REGION Network 10
   RUNG wire#powerrail
      Contact( "EstadosCmpALTA-MTA"._4s1 )
      I_Contact( "CompALTA-MTA".ReqMch4 )
      wire#w1
      Contact( "DB-CompAltaDatos".Aut4 )
      Coil( "Concatenadoras"._4c10 )
   END_RUNG
   RUNG wire#powerrail
      Contact( "EstadosCmpALTA-MTA"._4s9 )
      I_Contact( "CompALTA-MTA".ReqMch4 )
   END_RUNG wire#w1
   RUNG wire#powerrail
      Contact( "EstadosCmpALTA-MTA"._4s3 )
      I_Contact( "DB-CompAltaDatos".PanMchCmp4 )
   END_RUNG wire#w1
   // the same network as SCL:
   "Concatenadoras"._4c10 := (("EstadosCmpALTA-MTA"._4s1 AND NOT "CompALTA-MTA".ReqMch4) OR ("EstadosCmpALTA-MTA"._4s9 AND NOT "CompALTA-MTA".ReqMch4) OR ("EstadosCmpALTA-MTA"._4s3 AND NOT "DB-CompAltaDatos".PanMchCmp4)) AND "DB-CompAltaDatos".Aut4;
END_REGION

REGION Network 11
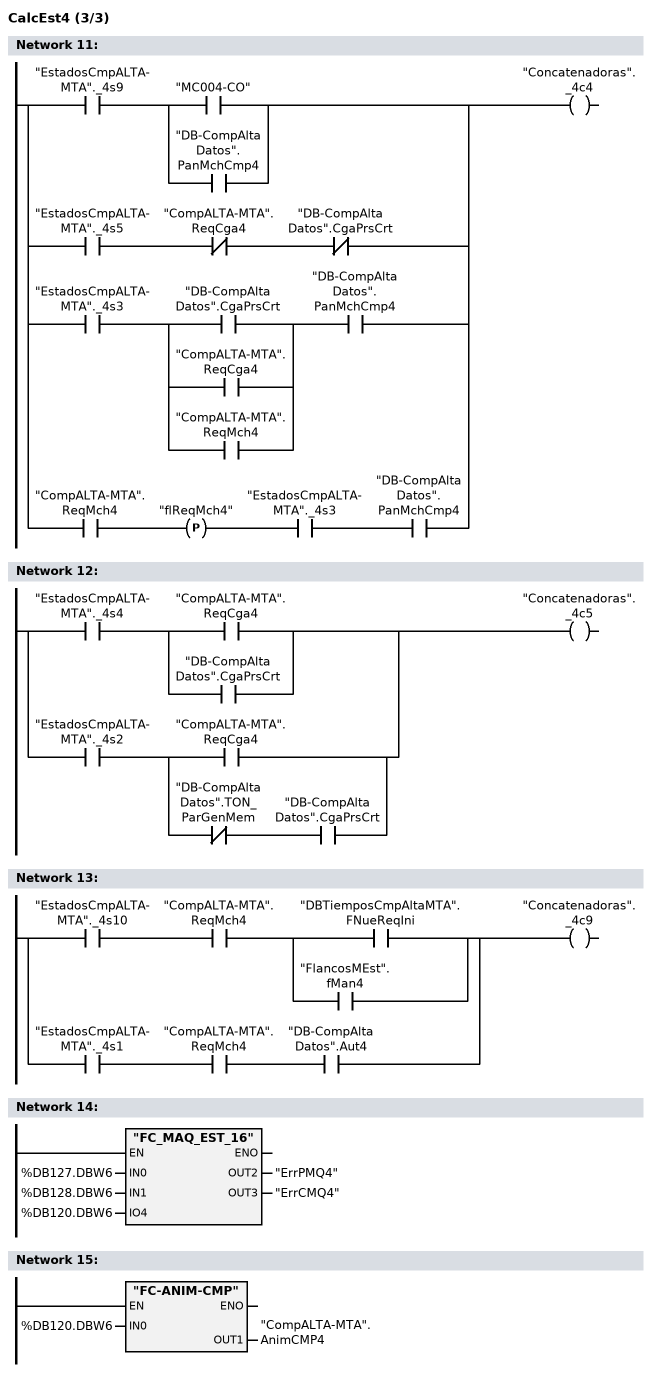
   RUNG wire#powerrail
      Contact( "EstadosCmpALTA-MTA"._4s9 )
      wire#w1
      Contact( "MC004-CO" )
      wire#w2
      Coil( "Concatenadoras"._4c4 )
   END_RUNG
   RUNG wire#w1
      Contact( "DB-CompAltaDatos".PanMchCmp4 )
   END_RUNG wire#w2
   RUNG wire#powerrail
      Contact( "EstadosCmpALTA-MTA"._4s5 )
      I_Contact( "CompALTA-MTA".ReqCga4 )
      I_Contact( "DB-CompAltaDatos".CgaPrsCrt )
   END_RUNG wire#w2
   RUNG wire#powerrail
      Contact( "EstadosCmpALTA-MTA"._4s3 )
      wire#w3
      Contact( "DB-CompAltaDatos".CgaPrsCrt )
      wire#w4
      Contact( "DB-CompAltaDatos".PanMchCmp4 )
   END_RUNG wire#w2
   RUNG wire#w3
      Contact( "CompALTA-MTA".ReqCga4 )
   END_RUNG wire#w4
   RUNG wire#w3
      Contact( "CompALTA-MTA".ReqMch4 )
   END_RUNG wire#w4
   RUNG wire#powerrail
      Contact( "CompALTA-MTA".ReqMch4 )
      P_Trig( "flReqMch4" )
      Contact( "EstadosCmpALTA-MTA"._4s3 )
      Contact( "DB-CompAltaDatos".PanMchCmp4 )
   END_RUNG wire#w2
   // the same network as SCL:
   #_w1 := "CompALTA-MTA".ReqMch4 AND NOT "flReqMch4";   // rising edge
   "flReqMch4" := "CompALTA-MTA".ReqMch4;
   "Concatenadoras"._4c4 := ("EstadosCmpALTA-MTA"._4s9 AND ("MC004-CO" OR "DB-CompAltaDatos".PanMchCmp4)) OR ("EstadosCmpALTA-MTA"._4s5 AND NOT "CompALTA-MTA".ReqCga4 AND NOT "DB-CompAltaDatos".CgaPrsCrt) OR ("EstadosCmpALTA-MTA"._4s3 AND ("DB-CompAltaDatos".CgaPrsCrt OR "CompALTA-MTA".ReqCga4 OR "CompALTA-MTA".ReqMch4) AND "DB-CompAltaDatos".PanMchCmp4) OR (#_w1 AND "EstadosCmpALTA-MTA"._4s3 AND "DB-CompAltaDatos".PanMchCmp4);
END_REGION

REGION Network 12
   RUNG wire#powerrail
      Contact( "EstadosCmpALTA-MTA"._4s4 )
      wire#w1
      Contact( "CompALTA-MTA".ReqCga4 )
      wire#w2
      Coil( "Concatenadoras"._4c5 )
   END_RUNG
   RUNG wire#w1
      Contact( "DB-CompAltaDatos".CgaPrsCrt )
   END_RUNG wire#w2
   RUNG wire#powerrail
      Contact( "EstadosCmpALTA-MTA"._4s2 )
      wire#w3
      Contact( "CompALTA-MTA".ReqCga4 )
   END_RUNG wire#w2
   RUNG wire#w3
      I_Contact( "DB-CompAltaDatos".TON_ParGenMem )
      Contact( "DB-CompAltaDatos".CgaPrsCrt )
   END_RUNG wire#w2
   // the same network as SCL:
   "Concatenadoras"._4c5 := ("EstadosCmpALTA-MTA"._4s4 AND ("CompALTA-MTA".ReqCga4 OR "DB-CompAltaDatos".CgaPrsCrt)) OR ("EstadosCmpALTA-MTA"._4s2 AND ("CompALTA-MTA".ReqCga4 OR (NOT "DB-CompAltaDatos".TON_ParGenMem AND "DB-CompAltaDatos".CgaPrsCrt)));
END_REGION

REGION Network 13
   RUNG wire#powerrail
      Contact( "EstadosCmpALTA-MTA"._4s10 )
      Contact( "CompALTA-MTA".ReqMch4 )
      wire#w1
      Contact( "DBTiemposCmpAltaMTA".FNueReqIni )
      wire#w2
      Coil( "Concatenadoras"._4c9 )
   END_RUNG
   RUNG wire#w1
      Contact( "FlancosMEst".fMan4 )
   END_RUNG wire#w2
   RUNG wire#powerrail
      Contact( "EstadosCmpALTA-MTA"._4s1 )
      Contact( "CompALTA-MTA".ReqMch4 )
      Contact( "DB-CompAltaDatos".Aut4 )
   END_RUNG wire#w2
   // the same network as SCL:
   "Concatenadoras"._4c9 := ("EstadosCmpALTA-MTA"._4s10 AND "CompALTA-MTA".ReqMch4 AND ("DBTiemposCmpAltaMTA".FNueReqIni OR "FlancosMEst".fMan4)) OR ("EstadosCmpALTA-MTA"._4s1 AND "CompALTA-MTA".ReqMch4 AND "DB-CompAltaDatos".Aut4);
END_REGION

REGION Network 14
   RUNG wire#powerrail
      "FC_MAQ_EST_16"(IN0 := %DB127.DBW6, IN1 := %DB128.DBW6, IO4 := %DB120.DBW6, OUT2 => "ErrPMQ4", OUT3 => "ErrCMQ4")
   END_RUNG
   // the same network as SCL:
   "FC_MAQ_EST_16"(IN0 := %DB127.DBW6,
                   IN1 := %DB128.DBW6,
                   IO4 := %DB120.DBW6,
                   OUT2 => "ErrPMQ4",
                   OUT3 => "ErrCMQ4");
END_REGION

REGION Network 15
   RUNG wire#powerrail
      "FC-ANIM-CMP"(IN0 := %DB120.DBW6, OUT1 => "CompALTA-MTA".AnimCMP4)
   END_RUNG
   // the same network as SCL:
   "FC-ANIM-CMP"(IN0 := %DB120.DBW6, OUT1 => "CompALTA-MTA".AnimCMP4);
END_REGION
END_FUNCTION

FUNCTION "CalcEst5" : Void   // FC40, LAD
{ S7_Optimized_Access := 'FALSE' }
VERSION : 0.1
   VAR_TEMP   // added for the SCL form of the ladder/FBD networks
      _w1 : Bool;
   END_VAR
BEGIN

REGION Network 1: Prioritaria 1
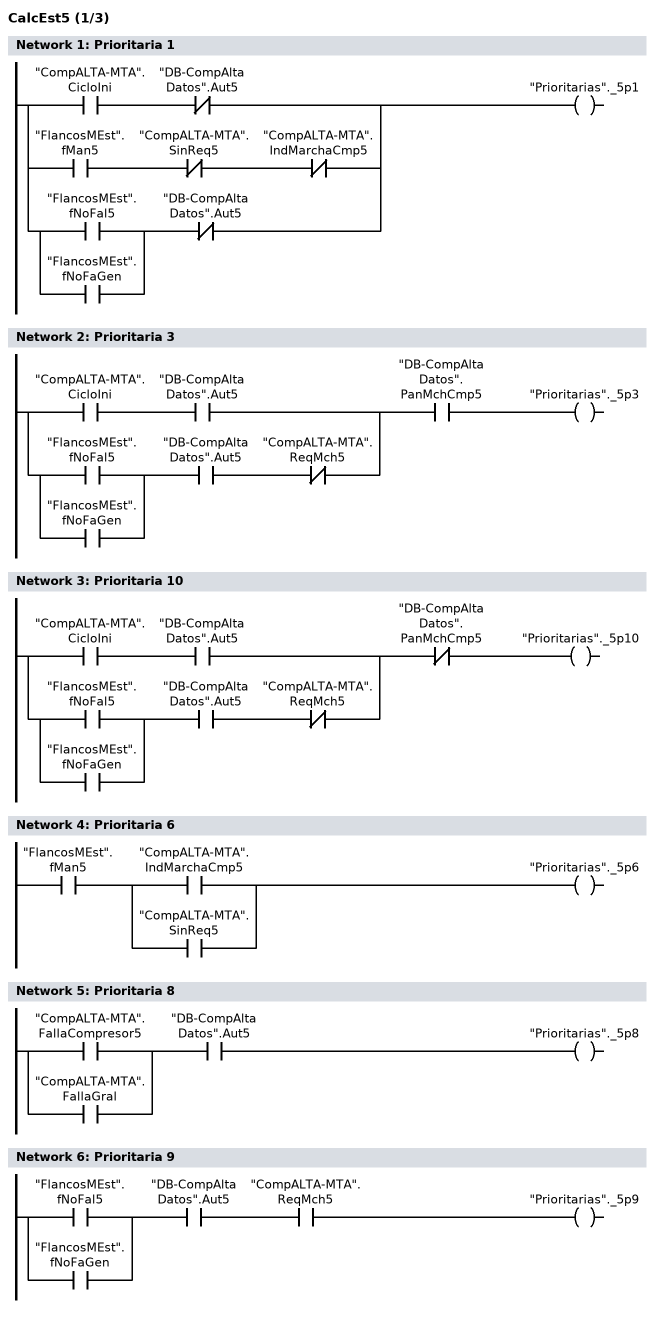
   RUNG wire#powerrail
      Contact( "CompALTA-MTA".CicloIni )
      I_Contact( "DB-CompAltaDatos".Aut5 )
      wire#w1
      Coil( "Prioritarias"._5p1 )
   END_RUNG
   RUNG wire#powerrail
      Contact( "FlancosMEst".fMan5 )
      I_Contact( "CompALTA-MTA".SinReq5 )
      I_Contact( "CompALTA-MTA".IndMarchaCmp5 )
   END_RUNG wire#w1
   RUNG wire#powerrail
      Contact( "FlancosMEst".fNoFal5 )
      wire#w2
      I_Contact( "DB-CompAltaDatos".Aut5 )
   END_RUNG wire#w1
   RUNG wire#powerrail
      Contact( "FlancosMEst".fNoFaGen )
   END_RUNG wire#w2
   // the same network as SCL:
   "Prioritarias"._5p1 := ("CompALTA-MTA".CicloIni AND NOT "DB-CompAltaDatos".Aut5) OR ("FlancosMEst".fMan5 AND NOT "CompALTA-MTA".SinReq5 AND NOT "CompALTA-MTA".IndMarchaCmp5) OR (("FlancosMEst".fNoFal5 OR "FlancosMEst".fNoFaGen) AND NOT "DB-CompAltaDatos".Aut5);
END_REGION

REGION Network 2: Prioritaria 3
   RUNG wire#powerrail
      Contact( "CompALTA-MTA".CicloIni )
      Contact( "DB-CompAltaDatos".Aut5 )
      wire#w1
      Contact( "DB-CompAltaDatos".PanMchCmp5 )
      Coil( "Prioritarias"._5p3 )
   END_RUNG
   RUNG wire#powerrail
      Contact( "FlancosMEst".fNoFal5 )
      wire#w2
      Contact( "DB-CompAltaDatos".Aut5 )
      I_Contact( "CompALTA-MTA".ReqMch5 )
   END_RUNG wire#w1
   RUNG wire#powerrail
      Contact( "FlancosMEst".fNoFaGen )
   END_RUNG wire#w2
   // the same network as SCL:
   "Prioritarias"._5p3 := (("CompALTA-MTA".CicloIni AND "DB-CompAltaDatos".Aut5) OR (("FlancosMEst".fNoFal5 OR "FlancosMEst".fNoFaGen) AND "DB-CompAltaDatos".Aut5 AND NOT "CompALTA-MTA".ReqMch5)) AND "DB-CompAltaDatos".PanMchCmp5;
END_REGION

REGION Network 3: Prioritaria 10
   RUNG wire#powerrail
      Contact( "CompALTA-MTA".CicloIni )
      Contact( "DB-CompAltaDatos".Aut5 )
      wire#w1
      I_Contact( "DB-CompAltaDatos".PanMchCmp5 )
      Coil( "Prioritarias"._5p10 )
   END_RUNG
   RUNG wire#powerrail
      Contact( "FlancosMEst".fNoFal5 )
      wire#w2
      Contact( "DB-CompAltaDatos".Aut5 )
      I_Contact( "CompALTA-MTA".ReqMch5 )
   END_RUNG wire#w1
   RUNG wire#powerrail
      Contact( "FlancosMEst".fNoFaGen )
   END_RUNG wire#w2
   // the same network as SCL:
   "Prioritarias"._5p10 := (("CompALTA-MTA".CicloIni AND "DB-CompAltaDatos".Aut5) OR (("FlancosMEst".fNoFal5 OR "FlancosMEst".fNoFaGen) AND "DB-CompAltaDatos".Aut5 AND NOT "CompALTA-MTA".ReqMch5)) AND NOT "DB-CompAltaDatos".PanMchCmp5;
END_REGION

REGION Network 4: Prioritaria 6
   RUNG wire#powerrail
      Contact( "FlancosMEst".fMan5 )
      wire#w1
      Contact( "CompALTA-MTA".IndMarchaCmp5 )
      wire#w2
      Coil( "Prioritarias"._5p6 )
   END_RUNG
   RUNG wire#w1
      Contact( "CompALTA-MTA".SinReq5 )
   END_RUNG wire#w2
   // the same network as SCL:
   "Prioritarias"._5p6 := "FlancosMEst".fMan5 AND ("CompALTA-MTA".IndMarchaCmp5 OR "CompALTA-MTA".SinReq5);
END_REGION

REGION Network 5: Prioritaria 8
   RUNG wire#powerrail
      Contact( "CompALTA-MTA".FallaCompresor5 )
      wire#w1
      Contact( "DB-CompAltaDatos".Aut5 )
      Coil( "Prioritarias"._5p8 )
   END_RUNG
   RUNG wire#powerrail
      Contact( "CompALTA-MTA".FallaGral )
   END_RUNG wire#w1
   // the same network as SCL:
   "Prioritarias"._5p8 := ("CompALTA-MTA".FallaCompresor5 OR "CompALTA-MTA".FallaGral) AND "DB-CompAltaDatos".Aut5;
END_REGION

REGION Network 6: Prioritaria 9
   RUNG wire#powerrail
      Contact( "FlancosMEst".fNoFal5 )
      wire#w1
      Contact( "DB-CompAltaDatos".Aut5 )
      Contact( "CompALTA-MTA".ReqMch5 )
      Coil( "Prioritarias"._5p9 )
   END_RUNG
   RUNG wire#powerrail
      Contact( "FlancosMEst".fNoFaGen )
   END_RUNG wire#w1
   // the same network as SCL:
   "Prioritarias"._5p9 := ("FlancosMEst".fNoFal5 OR "FlancosMEst".fNoFaGen) AND "DB-CompAltaDatos".Aut5 AND "CompALTA-MTA".ReqMch5;
END_REGION

REGION Network 7: Concatenadora 1
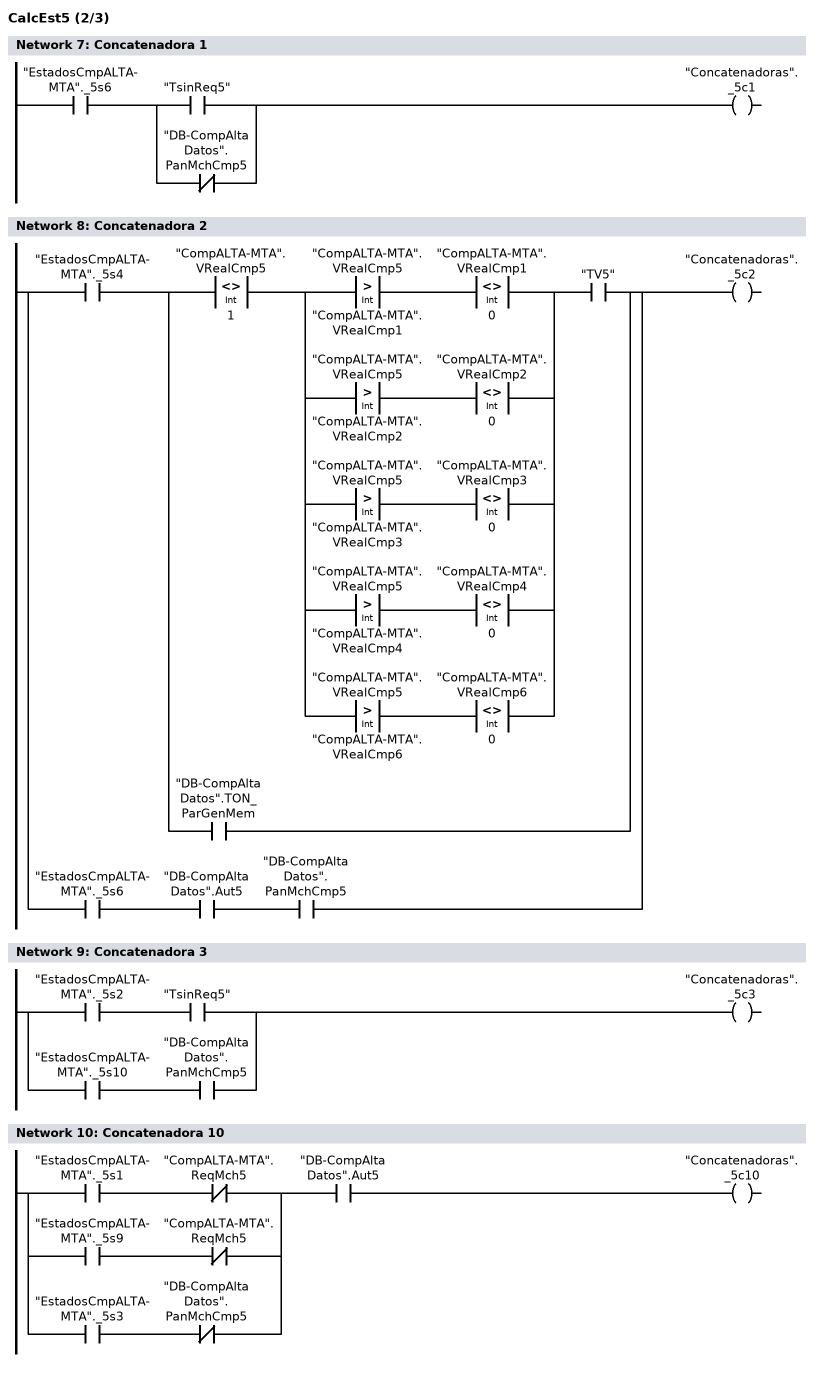
   RUNG wire#powerrail
      Contact( "EstadosCmpALTA-MTA"._5s6 )
      wire#w1
      Contact( "TsinReq5" )
      wire#w2
      Coil( "Concatenadoras"._5c1 )
   END_RUNG
   RUNG wire#w1
      I_Contact( "DB-CompAltaDatos".PanMchCmp5 )
   END_RUNG wire#w2
   // the same network as SCL:
   "Concatenadoras"._5c1 := "EstadosCmpALTA-MTA"._5s6 AND ("TsinReq5" OR NOT "DB-CompAltaDatos".PanMchCmp5);
END_REGION

REGION Network 8: Concatenadora 2
   RUNG wire#powerrail
      Contact( "EstadosCmpALTA-MTA"._5s4 )
      wire#w1
      { S7_Templates := "SrcType := Int" } NE_Contact(in1 := "CompALTA-MTA".VRealCmp5, in2 := 1)
      wire#w2
      { S7_Templates := "SrcType := Int" } GT_Contact(in1 := "CompALTA-MTA".VRealCmp5, in2 := "CompALTA-MTA".VRealCmp1)
      { S7_Templates := "SrcType := Int" } NE_Contact(in1 := "CompALTA-MTA".VRealCmp1, in2 := 0)
      wire#w3
      Contact( "TV5" )
      wire#w4
      Coil( "Concatenadoras"._5c2 )
   END_RUNG
   RUNG wire#w2
      { S7_Templates := "SrcType := Int" } GT_Contact(in1 := "CompALTA-MTA".VRealCmp5, in2 := "CompALTA-MTA".VRealCmp2)
      { S7_Templates := "SrcType := Int" } NE_Contact(in1 := "CompALTA-MTA".VRealCmp2, in2 := 0)
   END_RUNG wire#w3
   RUNG wire#w2
      { S7_Templates := "SrcType := Int" } GT_Contact(in1 := "CompALTA-MTA".VRealCmp5, in2 := "CompALTA-MTA".VRealCmp3)
      { S7_Templates := "SrcType := Int" } NE_Contact(in1 := "CompALTA-MTA".VRealCmp3, in2 := 0)
   END_RUNG wire#w3
   RUNG wire#w2
      { S7_Templates := "SrcType := Int" } GT_Contact(in1 := "CompALTA-MTA".VRealCmp5, in2 := "CompALTA-MTA".VRealCmp4)
      { S7_Templates := "SrcType := Int" } NE_Contact(in1 := "CompALTA-MTA".VRealCmp4, in2 := 0)
   END_RUNG wire#w3
   RUNG wire#w2
      { S7_Templates := "SrcType := Int" } GT_Contact(in1 := "CompALTA-MTA".VRealCmp5, in2 := "CompALTA-MTA".VRealCmp6)
      { S7_Templates := "SrcType := Int" } NE_Contact(in1 := "CompALTA-MTA".VRealCmp6, in2 := 0)
   END_RUNG wire#w3
   RUNG wire#w1
      Contact( "DB-CompAltaDatos".TON_ParGenMem )
   END_RUNG wire#w4
   RUNG wire#powerrail
      Contact( "EstadosCmpALTA-MTA"._5s6 )
      Contact( "DB-CompAltaDatos".Aut5 )
      Contact( "DB-CompAltaDatos".PanMchCmp5 )
   END_RUNG wire#w4
   // the same network as SCL:
   "Concatenadoras"._5c2 := ("EstadosCmpALTA-MTA"._5s4 AND ((("CompALTA-MTA".VRealCmp5 <> 1) AND ((("CompALTA-MTA".VRealCmp5 > "CompALTA-MTA".VRealCmp1) AND ("CompALTA-MTA".VRealCmp1 <> 0)) OR (("CompALTA-MTA".VRealCmp5 > "CompALTA-MTA".VRealCmp2) AND ("CompALTA-MTA".VRealCmp2 <> 0)) OR (("CompALTA-MTA".VRealCmp5 > "CompALTA-MTA".VRealCmp3) AND ("CompALTA-MTA".VRealCmp3 <> 0)) OR (("CompALTA-MTA".VRealCmp5 > "CompALTA-MTA".VRealCmp4) AND ("CompALTA-MTA".VRealCmp4 <> 0)) OR (("CompALTA-MTA".VRealCmp5 > "CompALTA-MTA".VRealCmp6) AND ("CompALTA-MTA".VRealCmp6 <> 0))) AND "TV5") OR "DB-CompAltaDatos".TON_ParGenMem)) OR ("EstadosCmpALTA-MTA"._5s6 AND "DB-CompAltaDatos".Aut5 AND "DB-CompAltaDatos".PanMchCmp5);
END_REGION

REGION Network 9: Concatenadora 3
   RUNG wire#powerrail
      Contact( "EstadosCmpALTA-MTA"._5s2 )
      Contact( "TsinReq5" )
      wire#w1
      Coil( "Concatenadoras"._5c3 )
   END_RUNG
   RUNG wire#powerrail
      Contact( "EstadosCmpALTA-MTA"._5s10 )
      Contact( "DB-CompAltaDatos".PanMchCmp5 )
   END_RUNG wire#w1
   // the same network as SCL:
   "Concatenadoras"._5c3 := ("EstadosCmpALTA-MTA"._5s2 AND "TsinReq5") OR ("EstadosCmpALTA-MTA"._5s10 AND "DB-CompAltaDatos".PanMchCmp5);
END_REGION

REGION Network 10: Concatenadora 10
   RUNG wire#powerrail
      Contact( "EstadosCmpALTA-MTA"._5s1 )
      I_Contact( "CompALTA-MTA".ReqMch5 )
      wire#w1
      Contact( "DB-CompAltaDatos".Aut5 )
      Coil( "Concatenadoras"._5c10 )
   END_RUNG
   RUNG wire#powerrail
      Contact( "EstadosCmpALTA-MTA"._5s9 )
      I_Contact( "CompALTA-MTA".ReqMch5 )
   END_RUNG wire#w1
   RUNG wire#powerrail
      Contact( "EstadosCmpALTA-MTA"._5s3 )
      I_Contact( "DB-CompAltaDatos".PanMchCmp5 )
   END_RUNG wire#w1
   // the same network as SCL:
   "Concatenadoras"._5c10 := (("EstadosCmpALTA-MTA"._5s1 AND NOT "CompALTA-MTA".ReqMch5) OR ("EstadosCmpALTA-MTA"._5s9 AND NOT "CompALTA-MTA".ReqMch5) OR ("EstadosCmpALTA-MTA"._5s3 AND NOT "DB-CompAltaDatos".PanMchCmp5)) AND "DB-CompAltaDatos".Aut5;
END_REGION

REGION Network 11: Concatenadora 4
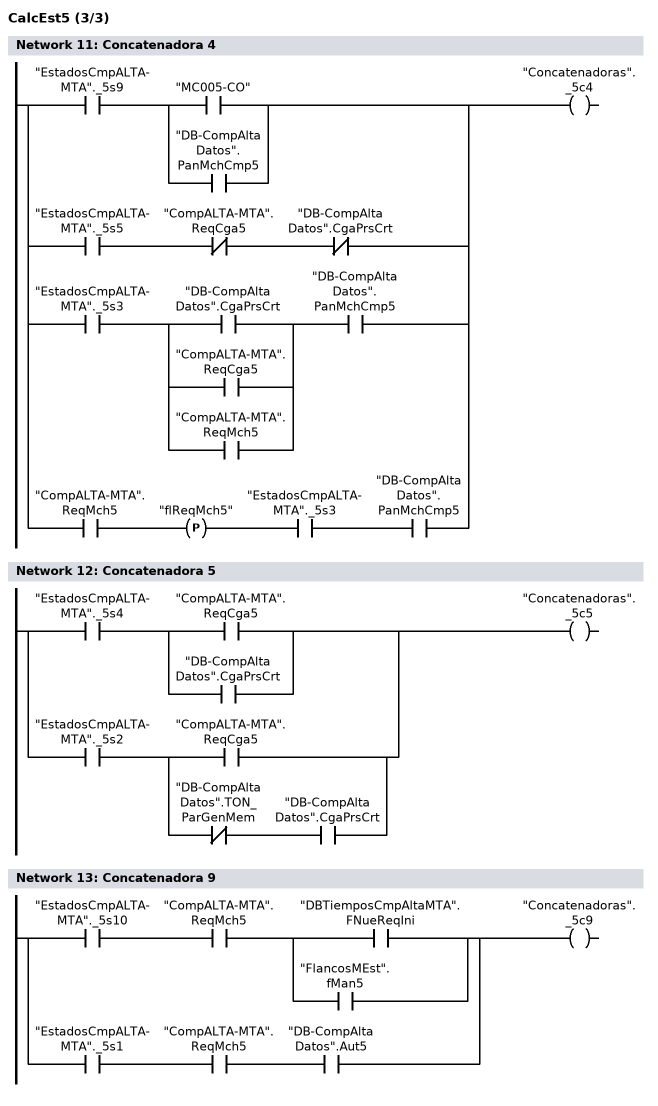
   RUNG wire#powerrail
      Contact( "EstadosCmpALTA-MTA"._5s9 )
      wire#w1
      Contact( "MC005-CO" )
      wire#w2
      Coil( "Concatenadoras"._5c4 )
   END_RUNG
   RUNG wire#w1
      Contact( "DB-CompAltaDatos".PanMchCmp5 )
   END_RUNG wire#w2
   RUNG wire#powerrail
      Contact( "EstadosCmpALTA-MTA"._5s5 )
      I_Contact( "CompALTA-MTA".ReqCga5 )
      I_Contact( "DB-CompAltaDatos".CgaPrsCrt )
   END_RUNG wire#w2
   RUNG wire#powerrail
      Contact( "EstadosCmpALTA-MTA"._5s3 )
      wire#w3
      Contact( "DB-CompAltaDatos".CgaPrsCrt )
      wire#w4
      Contact( "DB-CompAltaDatos".PanMchCmp5 )
   END_RUNG wire#w2
   RUNG wire#w3
      Contact( "CompALTA-MTA".ReqCga5 )
   END_RUNG wire#w4
   RUNG wire#w3
      Contact( "CompALTA-MTA".ReqMch5 )
   END_RUNG wire#w4
   RUNG wire#powerrail
      Contact( "CompALTA-MTA".ReqMch5 )
      P_Trig( "flReqMch5" )
      Contact( "EstadosCmpALTA-MTA"._5s3 )
      Contact( "DB-CompAltaDatos".PanMchCmp5 )
   END_RUNG wire#w2
   // the same network as SCL:
   #_w1 := "CompALTA-MTA".ReqMch5 AND NOT "flReqMch5";   // rising edge
   "flReqMch5" := "CompALTA-MTA".ReqMch5;
   "Concatenadoras"._5c4 := ("EstadosCmpALTA-MTA"._5s9 AND ("MC005-CO" OR "DB-CompAltaDatos".PanMchCmp5)) OR ("EstadosCmpALTA-MTA"._5s5 AND NOT "CompALTA-MTA".ReqCga5 AND NOT "DB-CompAltaDatos".CgaPrsCrt) OR ("EstadosCmpALTA-MTA"._5s3 AND ("DB-CompAltaDatos".CgaPrsCrt OR "CompALTA-MTA".ReqCga5 OR "CompALTA-MTA".ReqMch5) AND "DB-CompAltaDatos".PanMchCmp5) OR (#_w1 AND "EstadosCmpALTA-MTA"._5s3 AND "DB-CompAltaDatos".PanMchCmp5);
END_REGION

REGION Network 12: Concatenadora 5
   RUNG wire#powerrail
      Contact( "EstadosCmpALTA-MTA"._5s4 )
      wire#w1
      Contact( "CompALTA-MTA".ReqCga5 )
      wire#w2
      Coil( "Concatenadoras"._5c5 )
   END_RUNG
   RUNG wire#w1
      Contact( "DB-CompAltaDatos".CgaPrsCrt )
   END_RUNG wire#w2
   RUNG wire#powerrail
      Contact( "EstadosCmpALTA-MTA"._5s2 )
      wire#w3
      Contact( "CompALTA-MTA".ReqCga5 )
   END_RUNG wire#w2
   RUNG wire#w3
      I_Contact( "DB-CompAltaDatos".TON_ParGenMem )
      Contact( "DB-CompAltaDatos".CgaPrsCrt )
   END_RUNG wire#w2
   // the same network as SCL:
   "Concatenadoras"._5c5 := ("EstadosCmpALTA-MTA"._5s4 AND ("CompALTA-MTA".ReqCga5 OR "DB-CompAltaDatos".CgaPrsCrt)) OR ("EstadosCmpALTA-MTA"._5s2 AND ("CompALTA-MTA".ReqCga5 OR (NOT "DB-CompAltaDatos".TON_ParGenMem AND "DB-CompAltaDatos".CgaPrsCrt)));
END_REGION

REGION Network 13: Concatenadora 9
   RUNG wire#powerrail
      Contact( "EstadosCmpALTA-MTA"._5s10 )
      Contact( "CompALTA-MTA".ReqMch5 )
      wire#w1
      Contact( "DBTiemposCmpAltaMTA".FNueReqIni )
      wire#w2
      Coil( "Concatenadoras"._5c9 )
   END_RUNG
   RUNG wire#w1
      Contact( "FlancosMEst".fMan5 )
   END_RUNG wire#w2
   RUNG wire#powerrail
      Contact( "EstadosCmpALTA-MTA"._5s1 )
      Contact( "CompALTA-MTA".ReqMch5 )
      Contact( "DB-CompAltaDatos".Aut5 )
   END_RUNG wire#w2
   // the same network as SCL:
   "Concatenadoras"._5c9 := ("EstadosCmpALTA-MTA"._5s10 AND "CompALTA-MTA".ReqMch5 AND ("DBTiemposCmpAltaMTA".FNueReqIni OR "FlancosMEst".fMan5)) OR ("EstadosCmpALTA-MTA"._5s1 AND "CompALTA-MTA".ReqMch5 AND "DB-CompAltaDatos".Aut5);
END_REGION

REGION Network 14 (STL): Maquina de estados
         CALL  "FC_MAQ_EST_16"
         ( IN0  := %DB127.DBW8,
           IN1  := %DB128.DBW8,
           OUT2 := "ErrPMQ5",
           OUT3 := "ErrCMQ5",
           IO4  := %DB120.DBW8
         );
         NOP   0;
END_REGION

REGION Network 15 (STL): Bloque animación compresor
         CALL  "FC-ANIM-CMP"
         ( IN0  := %DB120.DBW8,
           OUT1 := "CompALTA-MTA".AnimCMP5
         );
         NOP   0;
END_REGION
END_FUNCTION

FUNCTION "CalcEst0" : Void   // FC42, LAD
{ S7_Optimized_Access := 'FALSE' }
VERSION : 0.1
BEGIN

REGION Network 1
